REGION Network 12: Output enabled M209 Fan
   RUNG wire#powerrail
      Contact( "Z201".ST_xCycleON )
      I_Contact( "DB_Z201_HMI".tAlm.tF.xM209FanFeedback )
      Coil( "Z201".ST_xOutputEnabledM209Chips )
   END_RUNG
   // the same network as SCL:
   "Z201".ST_xOutputEnabledM209Chips := "Z201".ST_xCycleON AND NOT "DB_Z201_HMI".tAlm.tF.xM209FanFeedback;
END_REGION

REGION Network 13: #### START/STOP ZONE ####
END_REGION

REGION Network 14: OS Start cycle
   RUNG wire#powerrail
      Contact( "DB_Z201_HMI".tHMW.xStartCycleRequest )
      wire#w1
      Coil( "Z201".OS_xStartCycle )
   END_RUNG
   RUNG wire#w1
      R_Coil( "DB_Z201_HMI".tHMW.xStartCycleRequest )
   END_RUNG
   // the same network as SCL:
   "Z201".OS_xStartCycle := "DB_Z201_HMI".tHMW.xStartCycleRequest;
   IF "DB_Z201_HMI".tHMW.xStartCycleRequest THEN "DB_Z201_HMI".tHMW.xStartCycleRequest := FALSE; END_IF;
END_REGION

REGION Network 15: OS Stop cycle
   RUNG wire#powerrail
      Contact( "DB_Z201_HMI".tHMW.xStopCycleRequest )
      wire#w1
      Coil( "Z201".OS_xStopCycle )
   END_RUNG
   RUNG wire#w1
      R_Coil( "DB_Z201_HMI".tHMW.xStopCycleRequest )
   END_RUNG
   // the same network as SCL:
   "Z201".OS_xStopCycle := "DB_Z201_HMI".tHMW.xStopCycleRequest;
   IF "DB_Z201_HMI".tHMW.xStopCycleRequest THEN "DB_Z201_HMI".tHMW.xStopCycleRequest := FALSE; END_IF;
END_REGION

REGION Network 16: OS Force stop cycle
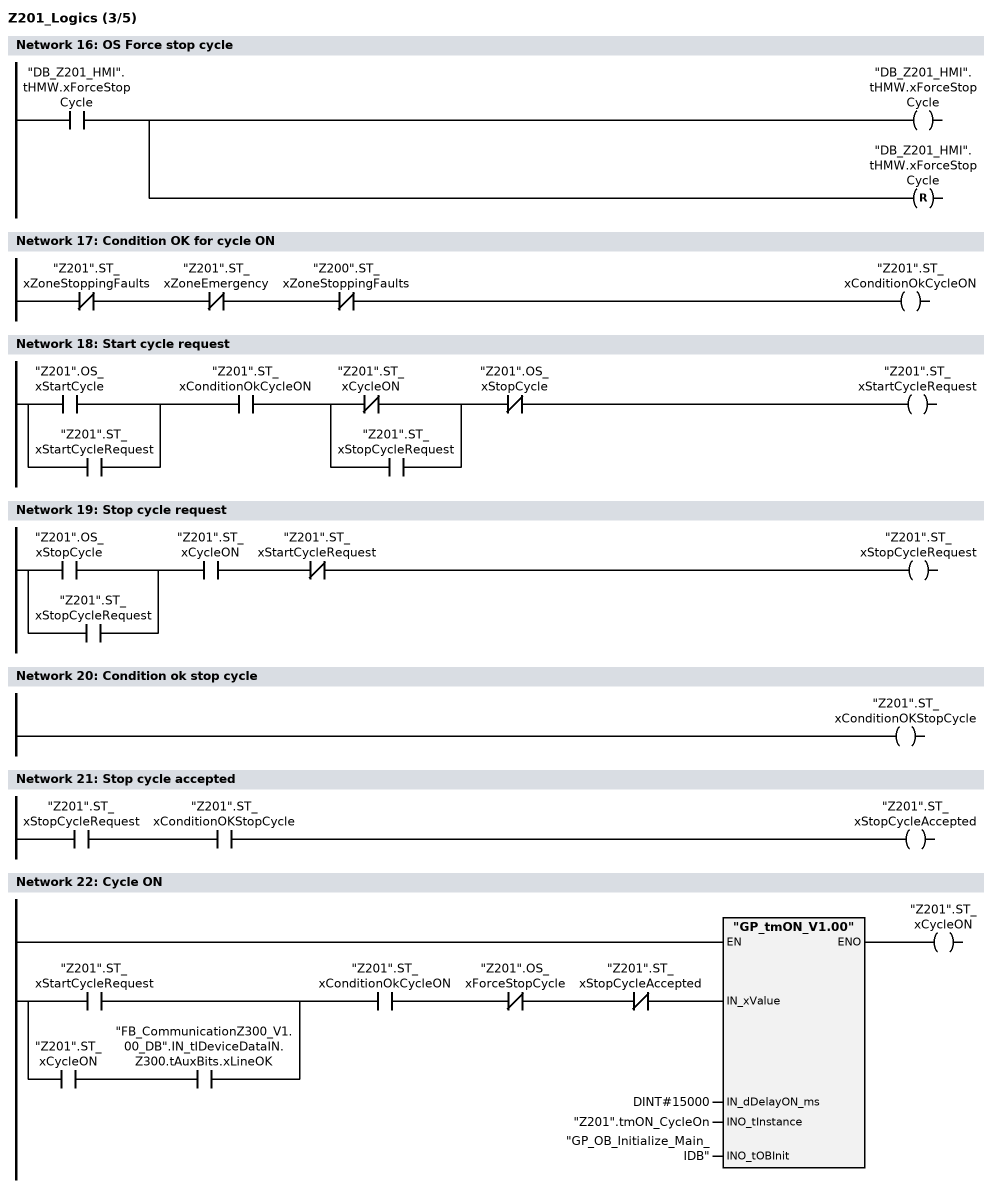
   RUNG wire#powerrail
      Contact( "DB_Z201_HMI".tHMW.xForceStopCycle )
      wire#w1
      Coil( "DB_Z201_HMI".tHMW.xForceStopCycle )
   END_RUNG
   RUNG wire#w1
      R_Coil( "DB_Z201_HMI".tHMW.xForceStopCycle )
   END_RUNG
   // the same network as SCL:
   #_w1 := "DB_Z201_HMI".tHMW.xForceStopCycle;
   "DB_Z201_HMI".tHMW.xForceStopCycle := "DB_Z201_HMI".tHMW.xForceStopCycle;
   IF #_w1 THEN "DB_Z201_HMI".tHMW.xForceStopCycle := FALSE; END_IF;
END_REGION

REGION Network 17: Condition OK for cycle ON
   RUNG wire#powerrail
      I_Contact( "Z201".ST_xZoneStoppingFaults )
      I_Contact( "Z201".ST_xZoneEmergency )
      I_Contact( "Z200".ST_xZoneStoppingFaults )
      Coil( "Z201".ST_xConditionOkCycleON )
   END_RUNG
   // the same network as SCL:
   "Z201".ST_xConditionOkCycleON := NOT "Z201".ST_xZoneStoppingFaults AND NOT "Z201".ST_xZoneEmergency AND NOT "Z200".ST_xZoneStoppingFaults;
END_REGION

REGION Network 18: Start cycle request
   RUNG wire#powerrail
      Contact( "Z201".OS_xStartCycle )
      wire#w1
      Contact( "Z201".ST_xConditionOkCycleON )
      wire#w2
      I_Contact( "Z201".ST_xCycleON )
      wire#w3
      I_Contact( "Z201".OS_xStopCycle )
      Coil( "Z201".ST_xStartCycleRequest )
   END_RUNG
   RUNG wire#powerrail
      Contact( "Z201".ST_xStartCycleRequest )
   END_RUNG wire#w1
   RUNG wire#w2
      Contact( "Z201".ST_xStopCycleRequest )
   END_RUNG wire#w3
   // the same network as SCL:
   "Z201".ST_xStartCycleRequest := ("Z201".OS_xStartCycle OR "Z201".ST_xStartCycleRequest) AND "Z201".ST_xConditionOkCycleON AND (NOT "Z201".ST_xCycleON OR "Z201".ST_xStopCycleRequest) AND NOT "Z201".OS_xStopCycle;
END_REGION

REGION Network 19: Stop cycle request
   RUNG wire#powerrail
      Contact( "Z201".OS_xStopCycle )
      wire#w1
      Contact( "Z201".ST_xCycleON )
      I_Contact( "Z201".ST_xStartCycleRequest )
      Coil( "Z201".ST_xStopCycleRequest )
   END_RUNG
   RUNG wire#powerrail
      Contact( "Z201".ST_xStopCycleRequest )
   END_RUNG wire#w1
   // the same network as SCL:
   "Z201".ST_xStopCycleRequest := ("Z201".OS_xStopCycle OR "Z201".ST_xStopCycleRequest) AND "Z201".ST_xCycleON AND NOT "Z201".ST_xStartCycleRequest;
END_REGION

REGION Network 20: Condition ok stop cycle
   RUNG wire#powerrail
      Coil( "Z201".ST_xConditionOKStopCycle )
   END_RUNG
   // the same network as SCL:
   "Z201".ST_xConditionOKStopCycle := TRUE;
END_REGION

REGION Network 21: Stop cycle accepted
   RUNG wire#powerrail
      Contact( "Z201".ST_xStopCycleRequest )
      Contact( "Z201".ST_xConditionOKStopCycle )
      Coil( "Z201".ST_xStopCycleAccepted )
   END_RUNG
   // the same network as SCL:
   "Z201".ST_xStopCycleAccepted := "Z201".ST_xStopCycleRequest AND "Z201".ST_xConditionOKStopCycle;
END_REGION

REGION Network 22: Cycle ON
   RUNG wire#powerrail
      "GP_tmON_V1.00"(IN_xValue := wire#w2, IN_dDelayON_ms := DINT#15000, INO_tInstance := "Z201".tmON_CycleOn, INO_tOBInit := "GP_OB_Initialize_Main_IDB")
      Coil( "Z201".ST_xCycleON )
   END_RUNG
   RUNG wire#powerrail
      Contact( "Z201".ST_xStartCycleRequest )
      wire#w1
      Contact( "Z201".ST_xConditionOkCycleON )
      I_Contact( "Z201".OS_xForceStopCycle )
      I_Contact( "Z201".ST_xStopCycleAccepted )
   END_RUNG wire#w2
   RUNG wire#powerrail
      Contact( "Z201".ST_xCycleON )
      Contact( "FB_CommunicationZ300_V1.00_DB".IN_tIDeviceDataIN.Z300.tAuxBits.xLineOK )
   END_RUNG wire#w1
   // the same network as SCL:
   "GP_tmON_V1.00"(IN_xValue := ("Z201".ST_xStartCycleRequest OR ("Z201".ST_xCycleON AND "FB_CommunicationZ300_V1.00_DB".IN_tIDeviceDataIN.Z300.tAuxBits.xLineOK)) AND "Z201".ST_xConditionOkCycleON AND NOT "Z201".OS_xForceStopCycle AND NOT "Z201".ST_xStopCycleAccepted,
                   IN_dDelayON_ms := DINT#15000,
                   INO_tInstance := "Z201".tmON_CycleOn,
                   INO_tOBInit := "GP_OB_Initialize_Main_IDB",
                   ENO => #_w1);
   "Z201".ST_xCycleON := #_w1;
END_REGION

REGION Network 23: Cycle ON delayed
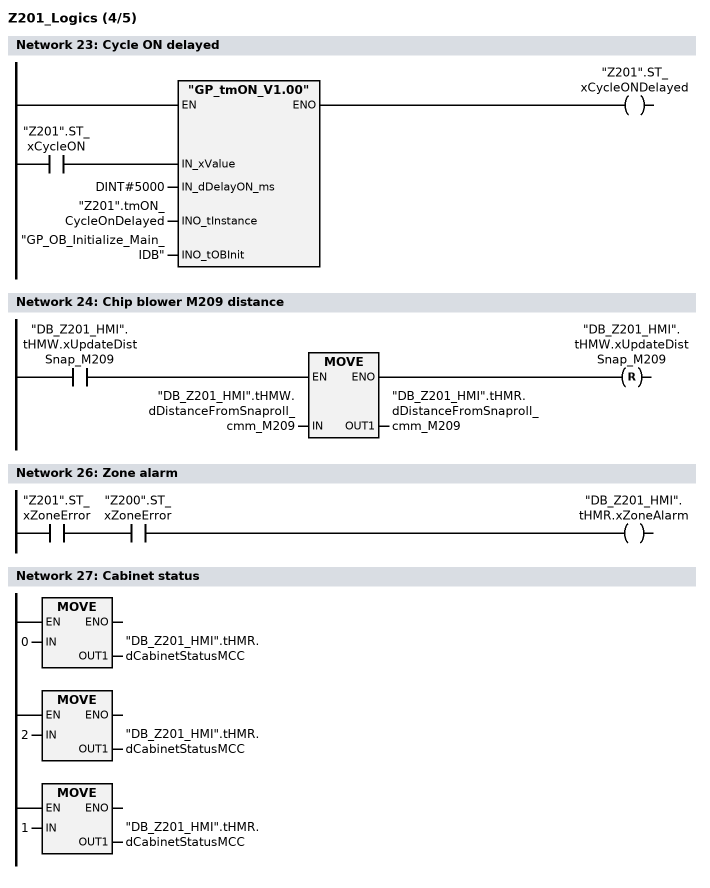
   RUNG wire#powerrail
      "GP_tmON_V1.00"(IN_xValue := wire#w1, IN_dDelayON_ms := DINT#5000, INO_tInstance := "Z201".tmON_CycleOnDelayed, INO_tOBInit := "GP_OB_Initialize_Main_IDB")
      Coil( "Z201".ST_xCycleONDelayed )
   END_RUNG
   RUNG wire#powerrail
      Contact( "Z201".ST_xCycleON )
   END_RUNG wire#w1
   // the same network as SCL:
   "GP_tmON_V1.00"(IN_xValue := "Z201".ST_xCycleON,
                   IN_dDelayON_ms := DINT#5000,
                   INO_tInstance := "Z201".tmON_CycleOnDelayed,
                   INO_tOBInit := "GP_OB_Initialize_Main_IDB",
                   ENO => #_w1);
   "Z201".ST_xCycleONDelayed := #_w1;
END_REGION

REGION Network 24: Chip blower M209 distance
   RUNG wire#powerrail
      Contact( "DB_Z201_HMI".tHMW.xUpdateDistSnap_M209 )
      Move(in := "DB_Z201_HMI".tHMW.dDistanceFromSnaproll_cmm_M209, out1 => "DB_Z201_HMI".tHMR.dDistanceFromSnaproll_cmm_M209)
      R_Coil( "DB_Z201_HMI".tHMW.xUpdateDistSnap_M209 )
   END_RUNG
   // the same network as SCL:
   IF "DB_Z201_HMI".tHMW.xUpdateDistSnap_M209 THEN
       "DB_Z201_HMI".tHMR.dDistanceFromSnaproll_cmm_M209 := "DB_Z201_HMI".tHMW.dDistanceFromSnaproll_cmm_M209;
       "DB_Z201_HMI".tHMW.xUpdateDistSnap_M209 := FALSE;
   END_IF;
END_REGION

REGION Network 25: #### HMI STATUSES ####
END_REGION

REGION Network 26: Zone alarm
   RUNG wire#powerrail
      Contact( "Z201".ST_xZoneError )
      Contact( "Z200".ST_xZoneError )
      Coil( "DB_Z201_HMI".tHMR.xZoneAlarm )
   END_RUNG
   // the same network as SCL:
   "DB_Z201_HMI".tHMR.xZoneAlarm := "Z201".ST_xZoneError AND "Z200".ST_xZoneError;
END_REGION

REGION Network 27: Cabinet status
   RUNG wire#powerrail
      Move(in := 0, out1 => "DB_Z201_HMI".tHMR.dCabinetStatusMCC)
   END_RUNG
   RUNG wire#powerrail
      Move(in := 2, out1 => "DB_Z201_HMI".tHMR.dCabinetStatusMCC)
   END_RUNG
   RUNG wire#powerrail
      Move(in := 1, out1 => "DB_Z201_HMI".tHMR.dCabinetStatusMCC)
   END_RUNG
   // the same network as SCL:
   "DB_Z201_HMI".tHMR.dCabinetStatusMCC := 0;
   "DB_Z201_HMI".tHMR.dCabinetStatusMCC := 2;
   "DB_Z201_HMI".tHMR.dCabinetStatusMCC := 1;
END_REGION

REGION Network 28: Zone state
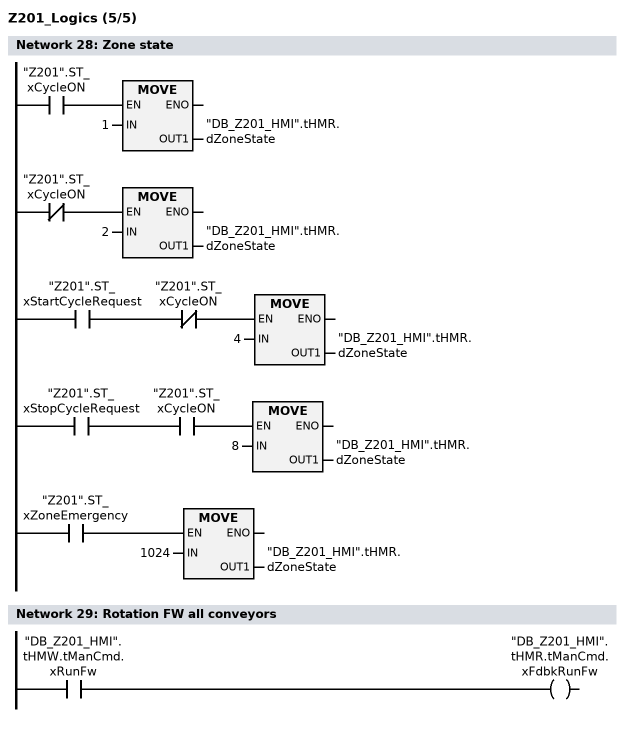
   RUNG wire#powerrail
      Contact( "Z201".ST_xCycleON )
      Move(in := 1, out1 => "DB_Z201_HMI".tHMR.dZoneState)
   END_RUNG
   RUNG wire#powerrail
      I_Contact( "Z201".ST_xCycleON )
      Move(in := 2, out1 => "DB_Z201_HMI".tHMR.dZoneState)
   END_RUNG
   RUNG wire#powerrail
      Contact( "Z201".ST_xStartCycleRequest )
      I_Contact( "Z201".ST_xCycleON )
      Move(in := 4, out1 => "DB_Z201_HMI".tHMR.dZoneState)
   END_RUNG
   RUNG wire#powerrail
      Contact( "Z201".ST_xStopCycleRequest )
      Contact( "Z201".ST_xCycleON )
      Move(in := 8, out1 => "DB_Z201_HMI".tHMR.dZoneState)
   END_RUNG
   RUNG wire#powerrail
      Contact( "Z201".ST_xZoneEmergency )
      Move(in := 1024, out1 => "DB_Z201_HMI".tHMR.dZoneState)
   END_RUNG
   // the same network as SCL:
   IF "Z201".ST_xCycleON THEN "DB_Z201_HMI".tHMR.dZoneState := 1; END_IF;
   IF NOT "Z201".ST_xCycleON THEN "DB_Z201_HMI".tHMR.dZoneState := 2; END_IF;
   IF "Z201".ST_xStartCycleRequest AND NOT "Z201".ST_xCycleON THEN
       "DB_Z201_HMI".tHMR.dZoneState := 4;
   END_IF;
   IF "Z201".ST_xStopCycleRequest AND "Z201".ST_xCycleON THEN "DB_Z201_HMI".tHMR.dZoneState := 8; END_IF;
   IF "Z201".ST_xZoneEmergency THEN "DB_Z201_HMI".tHMR.dZoneState := 1024; END_IF;
END_REGION

REGION Network 29: Rotation FW all conveyors
   RUNG wire#powerrail
      Contact( "DB_Z201_HMI".tHMW.tManCmd.xRunFw )
      Coil( "DB_Z201_HMI".tHMR.tManCmd.xFdbkRunFw )
   END_RUNG
   // the same network as SCL:
   "DB_Z201_HMI".tHMR.tManCmd.xFdbkRunFw := "DB_Z201_HMI".tHMW.tManCmd.xRunFw;
END_REGION

REGION Network 30: Enable/Disable Fan
   // Direttamente da scada
END_REGION
END_FUNCTION

FUNCTION "Z201_Output" : Void   // FC32, LAD
{ S7_Optimized_Access := 'TRUE' }
VERSION : 0.1
   VAR CONSTANT
      CONST_DBREAKDOWNOFF_CMM : DInt := 100000;   // Break downstream offset [mm/100]
      CONST_DBREAKUPOFF_CMM : DInt := 100000;   // Break upstream offset [mm/100]
   END_VAR
BEGIN

REGION Network 1: M216 Fan
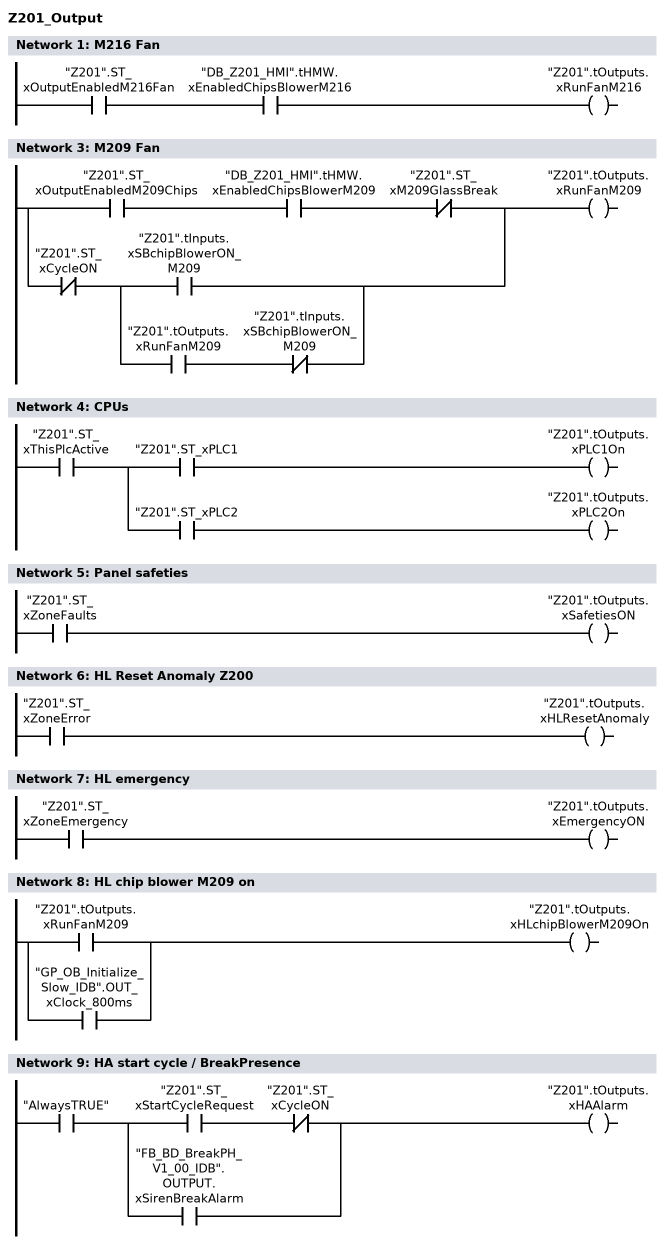
   RUNG wire#powerrail
      Contact( "Z201".ST_xOutputEnabledM216Fan )
      Contact( "DB_Z201_HMI".tHMW.xEnabledChipsBlowerM216 )
      Coil( "Z201".tOutputs.xRunFanM216 )
   END_RUNG
   // the same network as SCL:
   "Z201".tOutputs.xRunFanM216 := "Z201".ST_xOutputEnabledM216Fan AND "DB_Z201_HMI".tHMW.xEnabledChipsBlowerM216;
END_REGION

REGION Network 2 (SCL): Check glass break M209
   "DB_RibbonData".rgtGlassBreakRequest["DGLASSBREAKGET_M209"].IN_dDistanceSnaproll_cmm := "DB_Z201_HMI".tHMW.dDistanceFromSnaproll_cmm_M209;
   "DB_RibbonData".rgtGlassBreakRequest["DGLASSBREAKGET_M209"].IN_dDownstreamOffset_cmm := #CONST_DBREAKDOWNOFF_CMM;
   "DB_RibbonData".rgtGlassBreakRequest["DGLASSBREAKGET_M209"].IN_dUpstreamOffset_cmm := #CONST_DBREAKUPOFF_CMM;

   IF "DB_RibbonData".rgtGlassBreakRequest["DGLASSBREAKGET_M209"].OUT_xDataReady THEN
       "Z200".ST_xM209GlassBreak := "DB_RibbonData".rgtGlassBreakRequest["DGLASSBREAKGET_M209"].OUT_xGlassBreak;
   END_IF;

   IF "DB_RibbonData".rgtGlassBreakRequest["DGLASSBREAKGET_M209"].OUT_xDataReady OR NOT "DB_RibbonData".rgtGlassBreakRequest["DGLASSBREAKGET_M209"].IN_xRequestGlassBreak THEN
       "DB_RibbonData".rgtGlassBreakRequest["DGLASSBREAKGET_M209"].OUT_xDataReady := FALSE;
       "DB_RibbonData".rgtGlassBreakRequest["DGLASSBREAKGET_M209"].IN_xRequestGlassBreak := TRUE;
   END_IF;
END_REGION

REGION Network 3: M209 Fan
   RUNG wire#powerrail
      Contact( "Z201".ST_xOutputEnabledM209Chips )
      Contact( "DB_Z201_HMI".tHMW.xEnabledChipsBlowerM209 )
      I_Contact( "Z201".ST_xM209GlassBreak )
      wire#w1
      Coil( "Z201".tOutputs.xRunFanM209 )
   END_RUNG
   RUNG wire#powerrail
      I_Contact( "Z201".ST_xCycleON )
      wire#w2
      Contact( "Z201".tInputs.xSBchipBlowerON_M209 )
   END_RUNG wire#w1
   RUNG wire#w2
      Contact( "Z201".tOutputs.xRunFanM209 )
      I_Contact( "Z201".tInputs.xSBchipBlowerON_M209 )
   END_RUNG wire#w1
   // the same network as SCL:
   "Z201".tOutputs.xRunFanM209 := ("Z201".ST_xOutputEnabledM209Chips AND "DB_Z201_HMI".tHMW.xEnabledChipsBlowerM209 AND NOT "Z201".ST_xM209GlassBreak) OR (NOT "Z201".ST_xCycleON AND ("Z201".tInputs.xSBchipBlowerON_M209 OR ("Z201".tOutputs.xRunFanM209 AND NOT "Z201".tInputs.xSBchipBlowerON_M209)));
END_REGION

REGION Network 4: CPUs
   RUNG wire#powerrail
      Contact( "Z201".ST_xThisPlcActive )
      wire#w1
      Contact( "Z201".ST_xPLC1 )
      Coil( "Z201".tOutputs.xPLC1On )
   END_RUNG
   RUNG wire#w1
      Contact( "Z201".ST_xPLC2 )
      Coil( "Z201".tOutputs.xPLC2On )
   END_RUNG
   // the same network as SCL:
   "Z201".tOutputs.xPLC1On := "Z201".ST_xThisPlcActive AND "Z201".ST_xPLC1;
   "Z201".tOutputs.xPLC2On := "Z201".ST_xThisPlcActive AND "Z201".ST_xPLC2;
END_REGION

REGION Network 5: Panel safeties
   RUNG wire#powerrail
      Contact( "Z201".ST_xZoneFaults )
      Coil( "Z201".tOutputs.xSafetiesON )
   END_RUNG
   // the same network as SCL:
   "Z201".tOutputs.xSafetiesON := "Z201".ST_xZoneFaults;
END_REGION

REGION Network 6: HL Reset Anomaly Z200
   RUNG wire#powerrail
      Contact( "Z201".ST_xZoneError )
      Coil( "Z201".tOutputs.xHLResetAnomaly )
   END_RUNG
   // the same network as SCL:
   "Z201".tOutputs.xHLResetAnomaly := "Z201".ST_xZoneError;
END_REGION

REGION Network 7: HL emergency
   RUNG wire#powerrail
      Contact( "Z201".ST_xZoneEmergency )
      Coil( "Z201".tOutputs.xEmergencyON )
   END_RUNG
   // the same network as SCL:
   "Z201".tOutputs.xEmergencyON := "Z201".ST_xZoneEmergency;
END_REGION

REGION Network 8: HL chip blower M209 on
   RUNG wire#powerrail
      Contact( "Z201".tOutputs.xRunFanM209 )
      wire#w1
      Coil( "Z201".tOutputs.xHLchipBlowerM209On )
   END_RUNG
   RUNG wire#powerrail
      Contact( "GP_OB_Initialize_Slow_IDB".OUT_xClock_800ms )
   END_RUNG wire#w1
   // the same network as SCL:
   "Z201".tOutputs.xHLchipBlowerM209On := "Z201".tOutputs.xRunFanM209 OR "GP_OB_Initialize_Slow_IDB".OUT_xClock_800ms;
END_REGION

REGION Network 9: HA start cycle / BreakPresence
   RUNG wire#powerrail
      Contact( "AlwaysTRUE" )
      wire#w1
      Contact( "Z201".ST_xStartCycleRequest )
      I_Contact( "Z201".ST_xCycleON )
      wire#w2
      Coil( "Z201".tOutputs.xHAAlarm )
   END_RUNG
   RUNG wire#w1
      Contact( "FB_BD_BreakPH_V1_00_IDB".OUTPUT.xSirenBreakAlarm )
   END_RUNG wire#w2
   // the same network as SCL:
   "Z201".tOutputs.xHAAlarm := "AlwaysTRUE" AND (("Z201".ST_xStartCycleRequest AND NOT "Z201".ST_xCycleON) OR "FB_BD_BreakPH_V1_00_IDB".OUTPUT.xSirenBreakAlarm);
END_REGION
END_FUNCTION

FUNCTION "Z201_Faults" : Void   // FC152, LAD
{ S7_Optimized_Access := 'TRUE' }
VERSION : 0.1
   VAR_TEMP
      TMP_dwValue : DWord;
   END_VAR
   VAR_TEMP   // added for the SCL form of the ladder/FBD networks
      _w1 : Bool;
      _w2 : Bool;
   END_VAR
BEGIN

REGION Network 1 (SCL): Reset alarms
   IF "Z201".tmOFF_ResetAlarm.OUT_xDone THEN

       #TMP_dwValue := 0;

       SCATTER(IN:=#TMP_dwValue,
               OUT=>"DB_Z201_HMI".tAlm.tE);

       SCATTER(IN:=#TMP_dwValue,
               OUT=>"DB_Z201_HMI".tAlm.tS);

       SCATTER(IN:=#TMP_dwValue,
               OUT=>"DB_Z201_HMI".tAlm.tF);

       SCATTER(IN:=#TMP_dwValue,
               OUT=>"DB_Z201_HMI".tAlm.tW);

   END_IF;
END_REGION

REGION Network 2: ### EMERGENCY ###
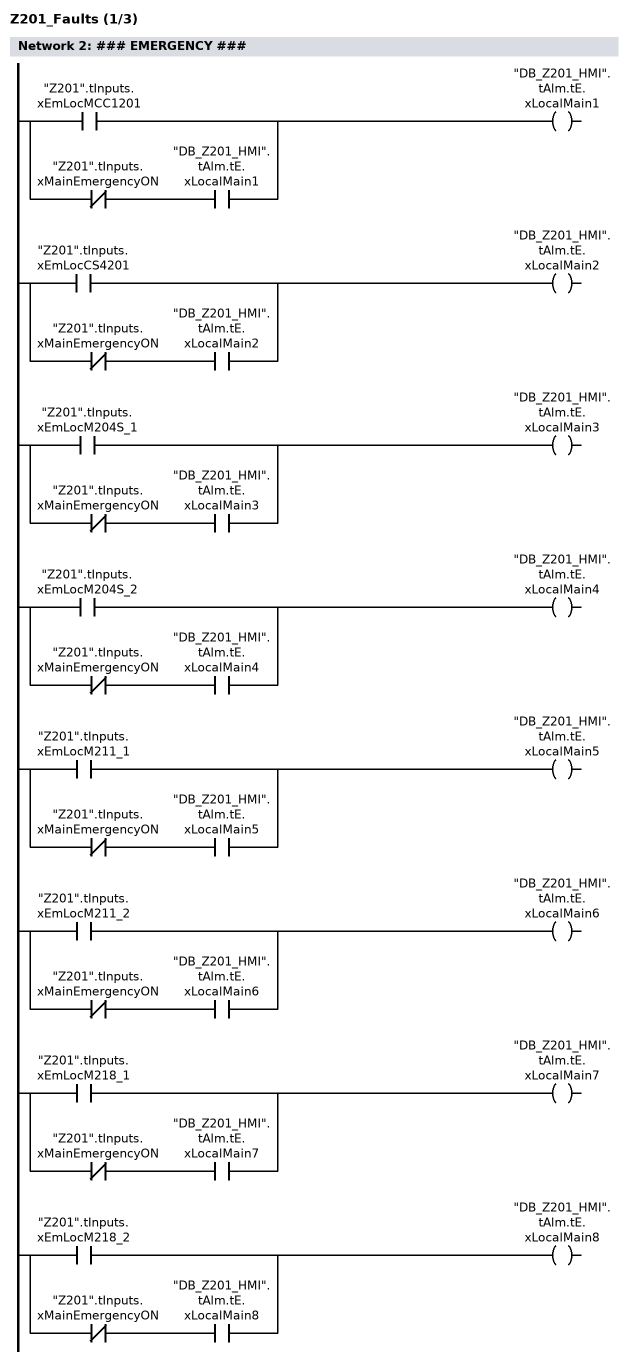
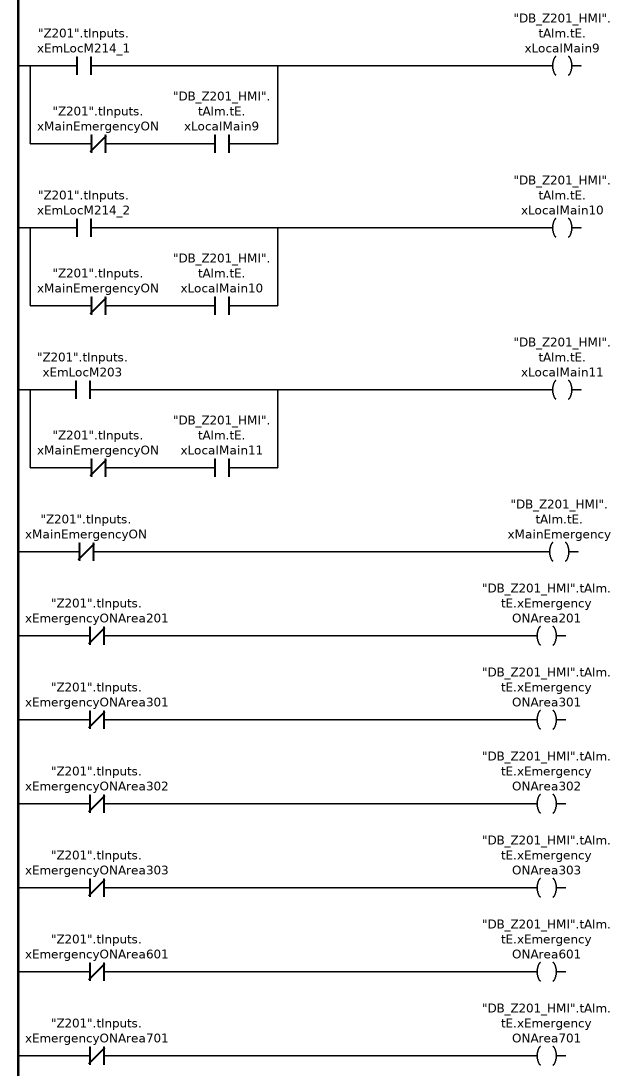
   RUNG wire#powerrail
      Contact( "Z201".tInputs.xEmLocMCC1201 )
      wire#w1
      Coil( "DB_Z201_HMI".tAlm.tE.xLocalMain1 )
   END_RUNG
   RUNG wire#powerrail
      I_Contact( "Z201".tInputs.xMainEmergencyON )
      Contact( "DB_Z201_HMI".tAlm.tE.xLocalMain1 )
   END_RUNG wire#w1
   RUNG wire#powerrail
      Contact( "Z201".tInputs.xEmLocCS4201 )
      wire#w2
      Coil( "DB_Z201_HMI".tAlm.tE.xLocalMain2 )
   END_RUNG
   RUNG wire#powerrail
      I_Contact( "Z201".tInputs.xMainEmergencyON )
      Contact( "DB_Z201_HMI".tAlm.tE.xLocalMain2 )
   END_RUNG wire#w2
   RUNG wire#powerrail
      Contact( "Z201".tInputs.xEmLocM204S_1 )
      wire#w3
      Coil( "DB_Z201_HMI".tAlm.tE.xLocalMain3 )
   END_RUNG
   RUNG wire#powerrail
      I_Contact( "Z201".tInputs.xMainEmergencyON )
      Contact( "DB_Z201_HMI".tAlm.tE.xLocalMain3 )
   END_RUNG wire#w3
   RUNG wire#powerrail
      Contact( "Z201".tInputs.xEmLocM204S_2 )
      wire#w4
      Coil( "DB_Z201_HMI".tAlm.tE.xLocalMain4 )
   END_RUNG
   RUNG wire#powerrail
      I_Contact( "Z201".tInputs.xMainEmergencyON )
      Contact( "DB_Z201_HMI".tAlm.tE.xLocalMain4 )
   END_RUNG wire#w4
   RUNG wire#powerrail
      Contact( "Z201".tInputs.xEmLocM211_1 )
      wire#w5
      Coil( "DB_Z201_HMI".tAlm.tE.xLocalMain5 )
   END_RUNG
   RUNG wire#powerrail
      I_Contact( "Z201".tInputs.xMainEmergencyON )
      Contact( "DB_Z201_HMI".tAlm.tE.xLocalMain5 )
   END_RUNG wire#w5
   RUNG wire#powerrail
      Contact( "Z201".tInputs.xEmLocM211_2 )
      wire#w6
      Coil( "DB_Z201_HMI".tAlm.tE.xLocalMain6 )
   END_RUNG
   RUNG wire#powerrail
      I_Contact( "Z201".tInputs.xMainEmergencyON )
      Contact( "DB_Z201_HMI".tAlm.tE.xLocalMain6 )
   END_RUNG wire#w6
   RUNG wire#powerrail
      Contact( "Z201".tInputs.xEmLocM218_1 )
      wire#w7
      Coil( "DB_Z201_HMI".tAlm.tE.xLocalMain7 )
   END_RUNG
   RUNG wire#powerrail
      I_Contact( "Z201".tInputs.xMainEmergencyON )
      Contact( "DB_Z201_HMI".tAlm.tE.xLocalMain7 )
   END_RUNG wire#w7
   RUNG wire#powerrail
      Contact( "Z201".tInputs.xEmLocM218_2 )
      wire#w8
      Coil( "DB_Z201_HMI".tAlm.tE.xLocalMain8 )
   END_RUNG
   RUNG wire#powerrail
      I_Contact( "Z201".tInputs.xMainEmergencyON )
      Contact( "DB_Z201_HMI".tAlm.tE.xLocalMain8 )
   END_RUNG wire#w8
   RUNG wire#powerrail
      Contact( "Z201".tInputs.xEmLocM214_1 )
      wire#w9
      Coil( "DB_Z201_HMI".tAlm.tE.xLocalMain9 )
   END_RUNG
   RUNG wire#powerrail
      I_Contact( "Z201".tInputs.xMainEmergencyON )
      Contact( "DB_Z201_HMI".tAlm.tE.xLocalMain9 )
   END_RUNG wire#w9
   RUNG wire#powerrail
      Contact( "Z201".tInputs.xEmLocM214_2 )
      wire#w10
      Coil( "DB_Z201_HMI".tAlm.tE.xLocalMain10 )
   END_RUNG
   RUNG wire#powerrail
      I_Contact( "Z201".tInputs.xMainEmergencyON )
      Contact( "DB_Z201_HMI".tAlm.tE.xLocalMain10 )
   END_RUNG wire#w10
   RUNG wire#powerrail
      Contact( "Z201".tInputs.xEmLocM203 )
      wire#w11
      Coil( "DB_Z201_HMI".tAlm.tE.xLocalMain11 )
   END_RUNG
   RUNG wire#powerrail
      I_Contact( "Z201".tInputs.xMainEmergencyON )
      Contact( "DB_Z201_HMI".tAlm.tE.xLocalMain11 )
   END_RUNG wire#w11
   RUNG wire#powerrail
      I_Contact( "Z201".tInputs.xMainEmergencyON )
      Coil( "DB_Z201_HMI".tAlm.tE.xMainEmergency )
   END_RUNG
   RUNG wire#powerrail
      I_Contact( "Z201".tInputs.xEmergencyONArea201 )
      Coil( "DB_Z201_HMI".tAlm.tE.xEmergencyONArea201 )
   END_RUNG
   RUNG wire#powerrail
      I_Contact( "Z201".tInputs.xEmergencyONArea301 )
      Coil( "DB_Z201_HMI".tAlm.tE.xEmergencyONArea301 )
   END_RUNG
   RUNG wire#powerrail
      I_Contact( "Z201".tInputs.xEmergencyONArea302 )
      Coil( "DB_Z201_HMI".tAlm.tE.xEmergencyONArea302 )
   END_RUNG
   RUNG wire#powerrail
      I_Contact( "Z201".tInputs.xEmergencyONArea303 )
      Coil( "DB_Z201_HMI".tAlm.tE.xEmergencyONArea303 )
   END_RUNG
   RUNG wire#powerrail
      I_Contact( "Z201".tInputs.xEmergencyONArea601 )
      Coil( "DB_Z201_HMI".tAlm.tE.xEmergencyONArea601 )
   END_RUNG
   RUNG wire#powerrail
      I_Contact( "Z201".tInputs.xEmergencyONArea701 )
      Coil( "DB_Z201_HMI".tAlm.tE.xEmergencyONArea701 )
   END_RUNG
   // the same network as SCL:
   "DB_Z201_HMI".tAlm.tE.xLocalMain1 := "Z201".tInputs.xEmLocMCC1201 OR (NOT "Z201".tInputs.xMainEmergencyON AND "DB_Z201_HMI".tAlm.tE.xLocalMain1);
   "DB_Z201_HMI".tAlm.tE.xLocalMain2 := "Z201".tInputs.xEmLocCS4201 OR (NOT "Z201".tInputs.xMainEmergencyON AND "DB_Z201_HMI".tAlm.tE.xLocalMain2);
   "DB_Z201_HMI".tAlm.tE.xLocalMain3 := "Z201".tInputs.xEmLocM204S_1 OR (NOT "Z201".tInputs.xMainEmergencyON AND "DB_Z201_HMI".tAlm.tE.xLocalMain3);
   "DB_Z201_HMI".tAlm.tE.xLocalMain4 := "Z201".tInputs.xEmLocM204S_2 OR (NOT "Z201".tInputs.xMainEmergencyON AND "DB_Z201_HMI".tAlm.tE.xLocalMain4);
   "DB_Z201_HMI".tAlm.tE.xLocalMain5 := "Z201".tInputs.xEmLocM211_1 OR (NOT "Z201".tInputs.xMainEmergencyON AND "DB_Z201_HMI".tAlm.tE.xLocalMain5);
   "DB_Z201_HMI".tAlm.tE.xLocalMain6 := "Z201".tInputs.xEmLocM211_2 OR (NOT "Z201".tInputs.xMainEmergencyON AND "DB_Z201_HMI".tAlm.tE.xLocalMain6);
   "DB_Z201_HMI".tAlm.tE.xLocalMain7 := "Z201".tInputs.xEmLocM218_1 OR (NOT "Z201".tInputs.xMainEmergencyON AND "DB_Z201_HMI".tAlm.tE.xLocalMain7);
   "DB_Z201_HMI".tAlm.tE.xLocalMain8 := "Z201".tInputs.xEmLocM218_2 OR (NOT "Z201".tInputs.xMainEmergencyON AND "DB_Z201_HMI".tAlm.tE.xLocalMain8);
   "DB_Z201_HMI".tAlm.tE.xLocalMain9 := "Z201".tInputs.xEmLocM214_1 OR (NOT "Z201".tInputs.xMainEmergencyON AND "DB_Z201_HMI".tAlm.tE.xLocalMain9);
   "DB_Z201_HMI".tAlm.tE.xLocalMain10 := "Z201".tInputs.xEmLocM214_2 OR (NOT "Z201".tInputs.xMainEmergencyON AND "DB_Z201_HMI".tAlm.tE.xLocalMain10);
   "DB_Z201_HMI".tAlm.tE.xLocalMain11 := "Z201".tInputs.xEmLocM203 OR (NOT "Z201".tInputs.xMainEmergencyON AND "DB_Z201_HMI".tAlm.tE.xLocalMain11);
   "DB_Z201_HMI".tAlm.tE.xMainEmergency := NOT "Z201".tInputs.xMainEmergencyON;
   "DB_Z201_HMI".tAlm.tE.xEmergencyONArea201 := NOT "Z201".tInputs.xEmergencyONArea201;
   "DB_Z201_HMI".tAlm.tE.xEmergencyONArea301 := NOT "Z201".tInputs.xEmergencyONArea301;
   "DB_Z201_HMI".tAlm.tE.xEmergencyONArea302 := NOT "Z201".tInputs.xEmergencyONArea302;
   "DB_Z201_HMI".tAlm.tE.xEmergencyONArea303 := NOT "Z201".tInputs.xEmergencyONArea303;
   "DB_Z201_HMI".tAlm.tE.xEmergencyONArea601 := NOT "Z201".tInputs.xEmergencyONArea601;
   "DB_Z201_HMI".tAlm.tE.xEmergencyONArea701 := NOT "Z201".tInputs.xEmergencyONArea701;
END_REGION

REGION Network 3: ### STOPPING FAULTS ###
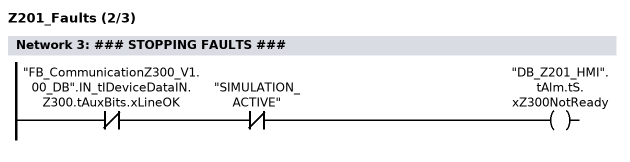
   RUNG wire#powerrail
      I_Contact( "FB_CommunicationZ300_V1.00_DB".IN_tIDeviceDataIN.Z300.tAuxBits.xLineOK )
      I_Contact( "SIMULATION_ACTIVE" )
      Coil( "DB_Z201_HMI".tAlm.tS.xZ300NotReady )
   END_RUNG
   // the same network as SCL:
   "DB_Z201_HMI".tAlm.tS.xZ300NotReady := NOT "FB_CommunicationZ300_V1.00_DB".IN_tIDeviceDataIN.Z300.tAuxBits.xLineOK AND NOT "SIMULATION_ACTIVE";
END_REGION

REGION Network 4: Anomalies / ### FAULTS ###
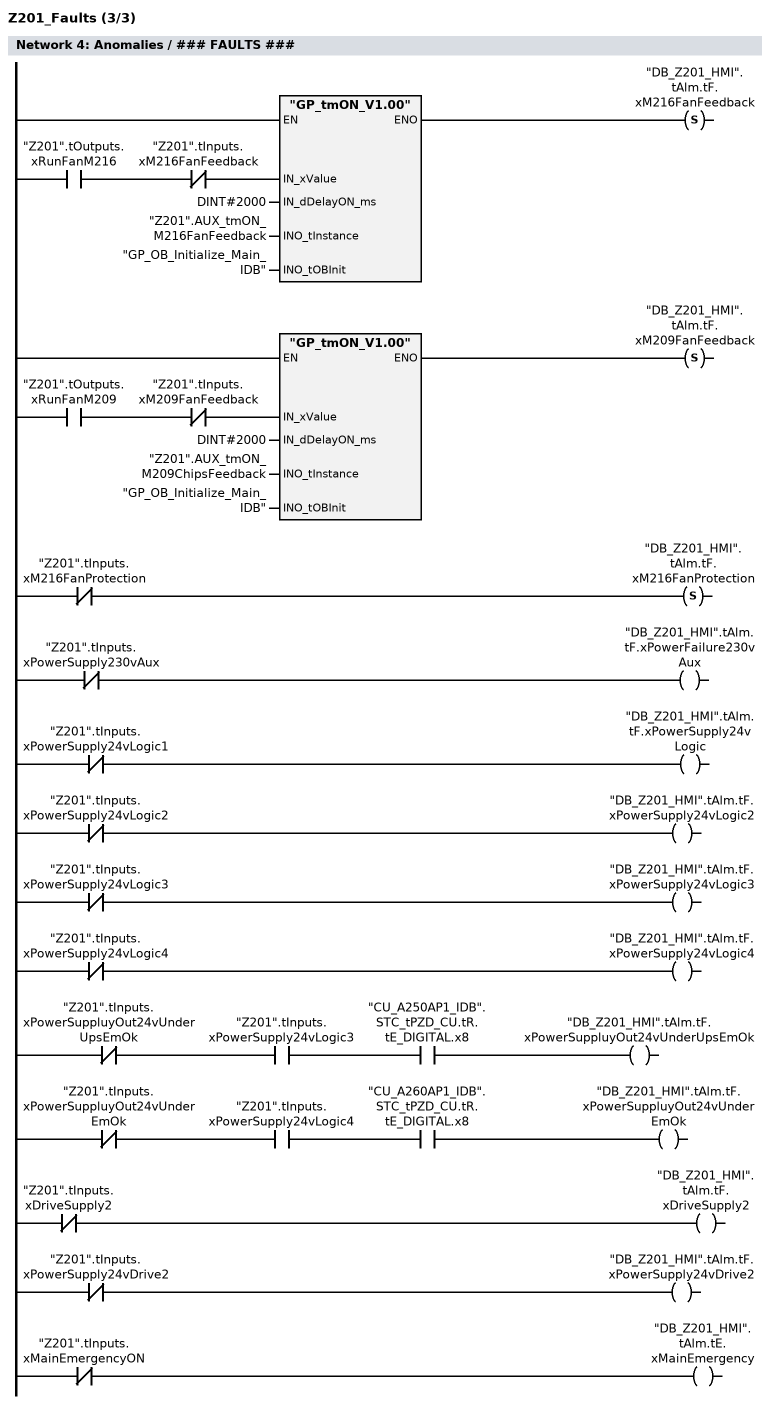
   RUNG wire#powerrail
      "GP_tmON_V1.00"(IN_xValue := wire#w1, IN_dDelayON_ms := DINT#2000, INO_tInstance := "Z201".AUX_tmON_M216FanFeedback, INO_tOBInit := "GP_OB_Initialize_Main_IDB")
      S_Coil( "DB_Z201_HMI".tAlm.tF.xM216FanFeedback )
   END_RUNG
   RUNG wire#powerrail
      Contact( "Z201".tOutputs.xRunFanM216 )
      I_Contact( "Z201".tInputs.xM216FanFeedback )
   END_RUNG wire#w1
   RUNG wire#powerrail
      "GP_tmON_V1.00"(IN_xValue := wire#w2, IN_dDelayON_ms := DINT#2000, INO_tInstance := "Z201".AUX_tmON_M209ChipsFeedback, INO_tOBInit := "GP_OB_Initialize_Main_IDB")
      S_Coil( "DB_Z201_HMI".tAlm.tF.xM209FanFeedback )
   END_RUNG
   RUNG wire#powerrail
      Contact( "Z201".tOutputs.xRunFanM209 )
      I_Contact( "Z201".tInputs.xM209FanFeedback )
   END_RUNG wire#w2
   RUNG wire#powerrail
      I_Contact( "Z201".tInputs.xM216FanProtection )
      S_Coil( "DB_Z201_HMI".tAlm.tF.xM216FanProtection )
   END_RUNG
   RUNG wire#powerrail
      I_Contact( "Z201".tInputs.xPowerSupply230vAux )
      Coil( "DB_Z201_HMI".tAlm.tF.xPowerFailure230vAux )
   END_RUNG
   RUNG wire#powerrail
      I_Contact( "Z201".tInputs.xPowerSupply24vLogic1 )
      Coil( "DB_Z201_HMI".tAlm.tF.xPowerSupply24vLogic )
   END_RUNG
   RUNG wire#powerrail
      I_Contact( "Z201".tInputs.xPowerSupply24vLogic2 )
      Coil( "DB_Z201_HMI".tAlm.tF.xPowerSupply24vLogic2 )
   END_RUNG
   RUNG wire#powerrail
      I_Contact( "Z201".tInputs.xPowerSupply24vLogic3 )
      Coil( "DB_Z201_HMI".tAlm.tF.xPowerSupply24vLogic3 )
   END_RUNG
   RUNG wire#powerrail
      I_Contact( "Z201".tInputs.xPowerSupply24vLogic4 )
      Coil( "DB_Z201_HMI".tAlm.tF.xPowerSupply24vLogic4 )
   END_RUNG
   RUNG wire#powerrail
      I_Contact( "Z201".tInputs.xPowerSuppluyOut24vUnderUpsEmOk )
      Contact( "Z201".tInputs.xPowerSupply24vLogic3 )
      Contact( "CU_A250AP1_IDB".STC_tPZD_CU.tR.tE_DIGITAL.x8 )
      Coil( "DB_Z201_HMI".tAlm.tF.xPowerSuppluyOut24vUnderUpsEmOk )
   END_RUNG
   RUNG wire#powerrail
      I_Contact( "Z201".tInputs.xPowerSuppluyOut24vUnderEmOk )
      Contact( "Z201".tInputs.xPowerSupply24vLogic4 )
      Contact( "CU_A260AP1_IDB".STC_tPZD_CU.tR.tE_DIGITAL.x8 )
      Coil( "DB_Z201_HMI".tAlm.tF.xPowerSuppluyOut24vUnderEmOk )
   END_RUNG
   RUNG wire#powerrail
      I_Contact( "Z201".tInputs.xDriveSupply2 )
      Coil( "DB_Z201_HMI".tAlm.tF.xDriveSupply2 )
   END_RUNG
   RUNG wire#powerrail
      I_Contact( "Z201".tInputs.xPowerSupply24vDrive2 )
      Coil( "DB_Z201_HMI".tAlm.tF.xPowerSupply24vDrive2 )
   END_RUNG
   RUNG wire#powerrail
      I_Contact( "Z201".tInputs.xMainEmergencyON )
      Coil( "DB_Z201_HMI".tAlm.tE.xMainEmergency )
   END_RUNG
   // the same network as SCL:
   "GP_tmON_V1.00"(IN_xValue := "Z201".tOutputs.xRunFanM216 AND NOT "Z201".tInputs.xM216FanFeedback,
                   IN_dDelayON_ms := DINT#2000,
                   INO_tInstance := "Z201".AUX_tmON_M216FanFeedback,
                   INO_tOBInit := "GP_OB_Initialize_Main_IDB",
                   ENO => #_w1);
   IF #_w1 THEN "DB_Z201_HMI".tAlm.tF.xM216FanFeedback := TRUE; END_IF;
   "GP_tmON_V1.00"(IN_xValue := "Z201".tOutputs.xRunFanM209 AND NOT "Z201".tInputs.xM209FanFeedback,
                   IN_dDelayON_ms := DINT#2000,
                   INO_tInstance := "Z201".AUX_tmON_M209ChipsFeedback,
                   INO_tOBInit := "GP_OB_Initialize_Main_IDB",
                   ENO => #_w2);
   IF #_w2 THEN "DB_Z201_HMI".tAlm.tF.xM209FanFeedback := TRUE; END_IF;
   IF NOT "Z201".tInputs.xM216FanProtection THEN "DB_Z201_HMI".tAlm.tF.xM216FanProtection := TRUE; END_IF;
   "DB_Z201_HMI".tAlm.tF.xPowerFailure230vAux := NOT "Z201".tInputs.xPowerSupply230vAux;
   "DB_Z201_HMI".tAlm.tF.xPowerSupply24vLogic := NOT "Z201".tInputs.xPowerSupply24vLogic1;
   "DB_Z201_HMI".tAlm.tF.xPowerSupply24vLogic2 := NOT "Z201".tInputs.xPowerSupply24vLogic2;
   "DB_Z201_HMI".tAlm.tF.xPowerSupply24vLogic3 := NOT "Z201".tInputs.xPowerSupply24vLogic3;
   "DB_Z201_HMI".tAlm.tF.xPowerSupply24vLogic4 := NOT "Z201".tInputs.xPowerSupply24vLogic4;
   "DB_Z201_HMI".tAlm.tF.xPowerSuppluyOut24vUnderUpsEmOk := NOT "Z201".tInputs.xPowerSuppluyOut24vUnderUpsEmOk AND "Z201".tInputs.xPowerSupply24vLogic3 AND "CU_A250AP1_IDB".STC_tPZD_CU.tR.tE_DIGITAL.x8;
   "DB_Z201_HMI".tAlm.tF.xPowerSuppluyOut24vUnderEmOk := NOT "Z201".tInputs.xPowerSuppluyOut24vUnderEmOk AND "Z201".tInputs.xPowerSupply24vLogic4 AND "CU_A260AP1_IDB".STC_tPZD_CU.tR.tE_DIGITAL.x8;
   "DB_Z201_HMI".tAlm.tF.xDriveSupply2 := NOT "Z201".tInputs.xDriveSupply2;
   "DB_Z201_HMI".tAlm.tF.xPowerSupply24vDrive2 := NOT "Z201".tInputs.xPowerSupply24vDrive2;
   "DB_Z201_HMI".tAlm.tE.xMainEmergency := NOT "Z201".tInputs.xMainEmergencyON;
END_REGION

REGION Network 5 (SCL): Calculate comulative status
   GATHER(IN:="DB_Z201_HMI".tAlm.tE,
              OUT=>#TMP_dwValue);

       IF "DB_Z201_HMI".tAlm.tE.xMainEmergency THEN
           "Z201".ST_xZoneEmergency := TRUE;
   ELSE
       "Z201".ST_xZoneEmergency := FALSE;
   END_IF;

   GATHER(IN:="DB_Z201_HMI".tAlm.tS,
              OUT=>#TMP_dwValue);

   IF #TMP_dwValue <> 0 THEN
       "Z201".ST_xZoneStoppingFaults := TRUE;
   ELSE
       "Z201".ST_xZoneStoppingFaults := FALSE;
   END_IF;

   GATHER(IN:="DB_Z201_HMI".tAlm.tF,
              OUT=>#TMP_dwValue);

   IF #TMP_dwValue <> 0 THEN
       "Z201".ST_xZoneFaults := TRUE;
   ELSE
       "Z201".ST_xZoneFaults := FALSE;
   END_IF;

   GATHER(IN:="DB_Z201_HMI".tAlm.tW,
              OUT=>#TMP_dwValue);

   IF #TMP_dwValue <> 0 THEN
       "Z201".ST_xZoneWarnings := TRUE;
   ELSE
       "Z201".ST_xZoneWarnings := FALSE;
   END_IF;

   IF "Z201".ST_xZoneEmergency AND "Z201".ST_xZoneStoppingFaults AND "Z201".ST_xZoneFaults THEN
       "Z201".ST_xZoneError := TRUE;
   ELSE
       "Z201".ST_xZoneError := FALSE;
   END_IF;
END_REGION
END_FUNCTION

// folder: 03_Programs_Logics/MCC1201/17_BreakDetector

